   "DB_Integer_S1AHour" : USInt = PLC Data_Integer.S1AHour, 1 s
   "DB_Integer_S1AMinute" : USInt = PLC Data_Integer.S1AMinute, 1 s
   "DB_Integer_S1ASecond" : USInt = PLC Data_Integer.S1ASecond, 1 s
   "DB_Integer_S1BHour" : USInt = PLC Data_Integer.S1BHour, 1 s
   "DB_Integer_S1BMinute" : USInt = PLC Data_Integer.S1BMinute, 1 s
   "DB_Integer_S1BSecond" : USInt = PLC Data_Integer.S1BSecond, 1 s
   "DB_Integer_S2AHour" : USInt = PLC Data_Integer.S2AHour, 1 s
   "DB_Integer_S2AMinute" : USInt = PLC Data_Integer.S2AMinute, 1 s
   "DB_Integer_S2ASecond" : USInt = PLC Data_Integer.S2ASecond, 1 s
   "DB_Integer_S2BHour" : USInt = PLC Data_Integer.S2BHour, 1 s
   "DB_Integer_S2BMinute" : USInt = PLC Data_Integer.S2BMinute, 1 s
   "DB_Integer_S2BSecond" : USInt = PLC Data_Integer.S2BSecond, 1 s
   "DB_Integer_S3AHour" : USInt = PLC Data_Integer.S3AHour, 1 s
   "DB_Integer_S3AMinute" : USInt = PLC Data_Integer.S3AMinute, 1 s
   "DB_Integer_S3ASecond" : USInt = PLC Data_Integer.S3ASecond, 1 s
   "DB_Integer_S3BHour" : USInt = PLC Data_Integer.S3BHour, 1 s
   "DB_Integer_S3BMinute" : USInt = PLC Data_Integer.S3BMinute, 1 s
   "DB_Integer_S3BSecond" : USInt = PLC Data_Integer.S3BSecond, 1 s
   "Data_Bool1_F_Set Time Day" : Bool = PLC Data_Bool1."F_Set Time Day", 1 s
   "Data_integer2_Flag Input Always Bad Read" : USInt = PLC Data_integer2."Flag Input Always Bad Read", 1 s
   "Data_DTLData_DTL_Mesin Run[0].HOUR" : USInt = PLC Data_DTLData."DTL_Mesin Run"[0].HOUR, 1 s
   "Data_DTLData_DTL_Mesin Run[0].MINUTE" : USInt = PLC Data_DTLData."DTL_Mesin Run"[0].MINUTE, 1 s
   "Data_DTLData_DTL_Mesin Run[0].SECOND" : USInt = PLC Data_DTLData."DTL_Mesin Run"[0].SECOND, 1 s
   "Data_Real_%Mesin Run[0]" : Real = PLC Data_Real."%Mesin Run"[0], 1 s
   "Data_DTLData_DTL_Mesin Run Baypass[0].HOUR" : USInt = PLC Data_DTLData."DTL_Mesin Run Baypass"[0].HOUR, 1 s
   "Data_DTLData_DTL_Mesin Run Baypass[0].MINUTE" : USInt = PLC Data_DTLData."DTL_Mesin Run Baypass"[0].MINUTE, 1 s
   "Data_DTLData_DTL_Mesin Run Baypass[0].SECOND" : USInt = PLC Data_DTLData."DTL_Mesin Run Baypass"[0].SECOND, 1 s
   "Data_Real_%Mesin Run Baypass[0]" : Real = PLC Data_Real."%Mesin Run Baypass"[0], 1 s
   "Data_DTLData_DTL_Mesin Stop[0].HOUR" : USInt = PLC Data_DTLData."DTL_Mesin Stop"[0].HOUR, 1 s
   "Data_DTLData_DTL_Mesin Stop[0].MINUTE" : USInt = PLC Data_DTLData."DTL_Mesin Stop"[0].MINUTE, 1 s
   "Data_DTLData_DTL_Mesin Stop[0].SECOND" : USInt = PLC Data_DTLData."DTL_Mesin Stop"[0].SECOND, 1 s
   "Data_Real_%Mesin Stop[0]" : Real = PLC Data_Real."%Mesin Stop"[0], 1 s
   "Data_DTLData_DTL_Mesin Error[0].HOUR" : USInt = PLC Data_DTLData."DTL_Mesin Error"[0].HOUR, 1 s
   "Data_DTLData_DTL_Mesin Error[0].MINUTE" : USInt = PLC Data_DTLData."DTL_Mesin Error"[0].MINUTE, 1 s
   "Data_DTLData_DTL_Mesin Error[0].SECOND" : USInt = PLC Data_DTLData."DTL_Mesin Error"[0].SECOND, 1 s
   "Data_Real_%Mesin Error[0]" : Real = PLC Data_Real."%Mesin Error"[0], 1 s
   "Data_DTLData_DTL_Mesin Run[1].HOUR" : USInt = PLC Data_DTLData."DTL_Mesin Run"[1].HOUR, 1 s
   "Data_DTLData_DTL_Mesin Run[1].MINUTE" : USInt = PLC Data_DTLData."DTL_Mesin Run"[1].MINUTE, 1 s
   "Data_DTLData_DTL_Mesin Run[1].SECOND" : USInt = PLC Data_DTLData."DTL_Mesin Run"[1].SECOND, 1 s
   "Data_Real_%Mesin Run[1]" : Real = PLC Data_Real."%Mesin Run"[1], 1 s
   "Data_DTLData_DTL_Mesin Run Baypass[1].HOUR" : USInt = PLC Data_DTLData."DTL_Mesin Run Baypass"[1].HOUR, 1 s
   "Data_DTLData_DTL_Mesin Run Baypass[1].MINUTE" : USInt = PLC Data_DTLData."DTL_Mesin Run Baypass"[1].MINUTE, 1 s
   "Data_DTLData_DTL_Mesin Run Baypass[1].SECOND" : USInt = PLC Data_DTLData."DTL_Mesin Run Baypass"[1].SECOND, 1 s
   "Data_Real_%Mesin Run Baypass[1]" : Real = PLC Data_Real."%Mesin Run Baypass"[1], 1 s
   "Data_DTLData_DTL_Mesin Stop[1].HOUR" : USInt = PLC Data_DTLData."DTL_Mesin Stop"[1].HOUR, 1 s
   "Data_DTLData_DTL_Mesin Stop[1].MINUTE" : USInt = PLC Data_DTLData."DTL_Mesin Stop"[1].MINUTE, 1 s
   "Data_DTLData_DTL_Mesin Stop[1].SECOND" : USInt = PLC Data_DTLData."DTL_Mesin Stop"[1].SECOND, 1 s
   "Data_Real_%Mesin Stop[1]" : Real = PLC Data_Real."%Mesin Stop"[1], 1 s
   "Data_DTLData_DTL_Mesin Error[1].HOUR" : USInt = PLC Data_DTLData."DTL_Mesin Error"[1].HOUR, 1 s
   "Data_DTLData_DTL_Mesin Error[1].MINUTE" : USInt = PLC Data_DTLData."DTL_Mesin Error"[1].MINUTE, 1 s
   "Data_DTLData_DTL_Mesin Error[1].SECOND" : USInt = PLC Data_DTLData."DTL_Mesin Error"[1].SECOND, 1 s
   "Data_Real_%Mesin Error[1]" : Real = PLC Data_Real."%Mesin Error"[1], 1 s
   "Data_DTLData_DTL_Mesin Run[2].HOUR" : USInt = PLC Data_DTLData."DTL_Mesin Run"[2].HOUR, 1 s
   "Data_DTLData_DTL_Mesin Run[2].MINUTE" : USInt = PLC Data_DTLData."DTL_Mesin Run"[2].MINUTE, 1 s
   "Data_DTLData_DTL_Mesin Run[2].SECOND" : USInt = PLC Data_DTLData."DTL_Mesin Run"[2].SECOND, 1 s
   "Data_Real_%Mesin Run[2]" : Real = PLC Data_Real."%Mesin Run"[2], 1 s
   "Data_DTLData_DTL_Mesin Run Baypass[2].HOUR" : USInt = PLC Data_DTLData."DTL_Mesin Run Baypass"[2].HOUR, 1 s
   "Data_DTLData_DTL_Mesin Run Baypass[2].MINUTE" : USInt = PLC Data_DTLData."DTL_Mesin Run Baypass"[2].MINUTE, 1 s
   "Data_DTLData_DTL_Mesin Run Baypass[2].SECOND" : USInt = PLC Data_DTLData."DTL_Mesin Run Baypass"[2].SECOND, 1 s
   "Data_Real_%Mesin Run Baypass[2]" : Real = PLC Data_Real."%Mesin Run Baypass"[2], 1 s
   "Data_DTLData_DTL_Mesin Stop[2].HOUR" : USInt = PLC Data_DTLData."DTL_Mesin Stop"[2].HOUR, 1 s
   "Data_DTLData_DTL_Mesin Stop[2].MINUTE" : USInt = PLC Data_DTLData."DTL_Mesin Stop"[2].MINUTE, 1 s
   "Data_DTLData_DTL_Mesin Stop[2].SECOND" : USInt = PLC Data_DTLData."DTL_Mesin Stop"[2].SECOND, 1 s
   "Data_Real_%Mesin Stop[2]" : Real = PLC Data_Real."%Mesin Stop"[2], 1 s
   "Data_DTLData_DTL_Mesin Error[2].HOUR" : USInt = PLC Data_DTLData."DTL_Mesin Error"[2].HOUR, 1 s
   "Data_DTLData_DTL_Mesin Error[2].MINUTE" : USInt = PLC Data_DTLData."DTL_Mesin Error"[2].MINUTE, 1 s
   "Data_DTLData_DTL_Mesin Error[2].SECOND" : USInt = PLC Data_DTLData."DTL_Mesin Error"[2].SECOND, 1 s
   "Data_Real_%Mesin Error[2]" : Real = PLC Data_Real."%Mesin Error"[2], 1 s
   "Data_DTLData_DTL_Mesin Run[3].HOUR" : USInt = PLC Data_DTLData."DTL_Mesin Run"[3].HOUR, 1 s
   "Data_DTLData_DTL_Mesin Run[3].MINUTE" : USInt = PLC Data_DTLData."DTL_Mesin Run"[3].MINUTE, 1 s
   "Data_DTLData_DTL_Mesin Run[3].SECOND" : USInt = PLC Data_DTLData."DTL_Mesin Run"[3].SECOND, 1 s
   "Data_Real_%Mesin Run[3]" : Real = PLC Data_Real."%Mesin Run"[3], 1 s
   "Data_DTLData_DTL_Mesin Run Baypass[3].HOUR" : USInt = PLC Data_DTLData."DTL_Mesin Run Baypass"[3].HOUR, 1 s
   "Data_DTLData_DTL_Mesin Run Baypass[3].MINUTE" : USInt = PLC Data_DTLData."DTL_Mesin Run Baypass"[3].MINUTE, 1 s
   "Data_DTLData_DTL_Mesin Run Baypass[3].SECOND" : USInt = PLC Data_DTLData."DTL_Mesin Run Baypass"[3].SECOND, 1 s
   "Data_Real_%Mesin Run Baypass[3]" : Real = PLC Data_Real."%Mesin Run Baypass"[3], 1 s
   "Data_Real_%Mesin Stop[3]" : Real = PLC Data_Real."%Mesin Stop"[3], 1 s
   "Data_Real_%Mesin Error[3]" : Real = PLC Data_Real."%Mesin Error"[3], 1 s
   "Data_DTLData_DTL_Mesin Stop[3].HOUR" : USInt = PLC Data_DTLData."DTL_Mesin Stop"[3].HOUR, 1 s
   "Data_DTLData_DTL_Mesin Stop[3].MINUTE" : USInt = PLC Data_DTLData."DTL_Mesin Stop"[3].MINUTE, 1 s
   "Data_DTLData_DTL_Mesin Stop[3].SECOND" : USInt = PLC Data_DTLData."DTL_Mesin Stop"[3].SECOND, 1 s
   "Data_DTLData_DTL_Mesin Error[3].HOUR" : USInt = PLC Data_DTLData."DTL_Mesin Error"[3].HOUR, 1 s
   "Data_DTLData_DTL_Mesin Error[3].MINUTE" : USInt = PLC Data_DTLData."DTL_Mesin Error"[3].MINUTE, 1 s
   "Data_DTLData_DTL_Mesin Error[3].SECOND" : USInt = PLC Data_DTLData."DTL_Mesin Error"[3].SECOND, 1 s
   "Data_DTLData_DTL_Mesin Run[4].HOUR" : USInt = PLC Data_DTLData."DTL_Mesin Run"[4].HOUR, 1 s
   "Data_DTLData_DTL_Mesin Run[4].MINUTE" : USInt = PLC Data_DTLData."DTL_Mesin Run"[4].MINUTE, 1 s
   "Data_DTLData_DTL_Mesin Run[4].SECOND" : USInt = PLC Data_DTLData."DTL_Mesin Run"[4].SECOND, 1 s
   "Data_Real_%Mesin Run[4]" : Real = PLC Data_Real."%Mesin Run"[4], 1 s
   "Data_Real_%Mesin Run Baypass[4]" : Real = PLC Data_Real."%Mesin Run Baypass"[4], 1 s
   "Data_Real_%Mesin Stop[4]" : Real = PLC Data_Real."%Mesin Stop"[4], 1 s
   "Data_Real_%Mesin Error[4]" : Real = PLC Data_Real."%Mesin Error"[4], 1 s
   "Data_DTLData_DTL_Mesin Run Baypass[4].HOUR" : USInt = PLC Data_DTLData."DTL_Mesin Run Baypass"[4].HOUR, 1 s
   "Data_DTLData_DTL_Mesin Run Baypass[4].MINUTE" : USInt = PLC Data_DTLData."DTL_Mesin Run Baypass"[4].MINUTE, 1 s
   "Data_DTLData_DTL_Mesin Run Baypass[4].SECOND" : USInt = PLC Data_DTLData."DTL_Mesin Run Baypass"[4].SECOND, 1 s
   "Data_DTLData_DTL_Mesin Stop[4].HOUR" : USInt = PLC Data_DTLData."DTL_Mesin Stop"[4].HOUR, 1 s
   "Data_DTLData_DTL_Mesin Stop[4].MINUTE" : USInt = PLC Data_DTLData."DTL_Mesin Stop"[4].MINUTE, 1 s
   "Data_DTLData_DTL_Mesin Stop[4].SECOND" : USInt = PLC Data_DTLData."DTL_Mesin Stop"[4].SECOND, 1 s
   "Data_DTLData_DTL_Mesin Error[4].HOUR" : USInt = PLC Data_DTLData."DTL_Mesin Error"[4].HOUR, 1 s
   "Data_DTLData_DTL_Mesin Error[4].MINUTE" : USInt = PLC Data_DTLData."DTL_Mesin Error"[4].MINUTE, 1 s
   "Data_DTLData_DTL_Mesin Error[4].SECOND" : USInt = PLC Data_DTLData."DTL_Mesin Error"[4].SECOND, 1 s
   "Data_DTLData_DTL_Mesin Run[5].HOUR" : USInt = PLC Data_DTLData."DTL_Mesin Run"[5].HOUR, 1 s
   "Data_DTLData_DTL_Mesin Run[5].MINUTE" : USInt = PLC Data_DTLData."DTL_Mesin Run"[5].MINUTE, 1 s
   "Data_DTLData_DTL_Mesin Run[5].SECOND" : USInt = PLC Data_DTLData."DTL_Mesin Run"[5].SECOND, 1 s
   "Data_Real_%Mesin Run[5]" : Real = PLC Data_Real."%Mesin Run"[5], 1 s
   "Data_Real_%Mesin Run Baypass[5]" : Real = PLC Data_Real."%Mesin Run Baypass"[5], 1 s
   "Data_Real_%Mesin Stop[5]" : Real = PLC Data_Real."%Mesin Stop"[5], 1 s
   "Data_Real_%Mesin Error[5]" : Real = PLC Data_Real."%Mesin Error"[5], 1 s
   "Data_DTLData_DTL_Mesin Run Baypass[5].HOUR" : USInt = PLC Data_DTLData."DTL_Mesin Run Baypass"[5].HOUR, 1 s
   "Data_DTLData_DTL_Mesin Run Baypass[5].MINUTE" : USInt = PLC Data_DTLData."DTL_Mesin Run Baypass"[5].MINUTE, 1 s
   "Data_DTLData_DTL_Mesin Run Baypass[5].SECOND" : USInt = PLC Data_DTLData."DTL_Mesin Run Baypass"[5].SECOND, 1 s
   "Data_DTLData_DTL_Mesin Stop[5].HOUR" : USInt = PLC Data_DTLData."DTL_Mesin Stop"[5].HOUR, 1 s
   "Data_DTLData_DTL_Mesin Stop[5].MINUTE" : USInt = PLC Data_DTLData."DTL_Mesin Stop"[5].MINUTE, 1 s
   "Data_DTLData_DTL_Mesin Stop[5].SECOND" : USInt = PLC Data_DTLData."DTL_Mesin Stop"[5].SECOND, 1 s
   "Data_DTLData_DTL_Mesin Error[5].HOUR" : USInt = PLC Data_DTLData."DTL_Mesin Error"[5].HOUR, 1 s
   "Data_DTLData_DTL_Mesin Error[5].MINUTE" : USInt = PLC Data_DTLData."DTL_Mesin Error"[5].MINUTE, 1 s
   "Data_DTLData_DTL_Mesin Error[5].SECOND" : USInt = PLC Data_DTLData."DTL_Mesin Error"[5].SECOND, 1 s
   "Data_Time_Timer Delay Stamp" : Time = PLC Data_Time."Timer Delay Stamp", 1 s
   "Data_Time_Timer Trigger Barcode" : Time = PLC Data_Time."Timer Trigger Barcode", 1 s
   "Data_Time_Timer Rejector Slof" : Time = PLC Data_Time."Timer Rejector Slof", 1 s
   "Data_Time_Timer AutoReject" : Time = PLC Data_Time."Timer AutoReject", 1 s
   "Data_DTLData_DTL_Always bad Read[0].HOUR" : USInt = PLC Data_DTLData."DTL_Always bad Read"[0].HOUR, 1 s
   "Data_DTLData_DTL_Always bad Read[0].MINUTE" : USInt = PLC Data_DTLData."DTL_Always bad Read"[0].MINUTE, 1 s
   "Data_DTLData_DTL_Always bad Read[0].SECOND" : USInt = PLC Data_DTLData."DTL_Always bad Read"[0].SECOND, 1 s
   "Data_DTLData_DTL_Press Low[0].HOUR" : USInt = PLC Data_DTLData."DTL_Press Low"[0].HOUR, 1 s
   "Data_DTLData_DTL_Press Low[0].MINUTE" : USInt = PLC Data_DTLData."DTL_Press Low"[0].MINUTE, 1 s
   "Data_DTLData_DTL_Press Low[0].SECOND" : USInt = PLC Data_DTLData."DTL_Press Low"[0].SECOND, 1 s
   "Data_DTLData_DTL_Door Open[0].HOUR" : USInt = PLC Data_DTLData."DTL_Door Open"[0].HOUR, 1 s
   "Data_DTLData_DTL_Door Open[0].MINUTE" : USInt = PLC Data_DTLData."DTL_Door Open"[0].MINUTE, 1 s
   "Data_DTLData_DTL_Door Open[0].SECOND" : USInt = PLC Data_DTLData."DTL_Door Open"[0].SECOND, 1 s
   "Data_DTLData_DTL_Total Detail Error[0].HOUR" : USInt = PLC Data_DTLData."DTL_Total Detail Error"[0].HOUR, 1 s
   "Data_DTLData_DTL_Total Detail Error[0].MINUTE" : USInt = PLC Data_DTLData."DTL_Total Detail Error"[0].MINUTE, 1 s
   "Data_DTLData_DTL_Total Detail Error[0].SECOND" : USInt = PLC Data_DTLData."DTL_Total Detail Error"[0].SECOND, 1 s
   "Data_DTLData_DTL_Always bad Read[1].HOUR" : USInt = PLC Data_DTLData."DTL_Always bad Read"[1].HOUR, 1 s
   "Data_DTLData_DTL_Always bad Read[1].MINUTE" : USInt = PLC Data_DTLData."DTL_Always bad Read"[1].MINUTE, 1 s
   "Data_DTLData_DTL_Always bad Read[1].SECOND" : USInt = PLC Data_DTLData."DTL_Always bad Read"[1].SECOND, 1 s
   "Data_DTLData_DTL_Press Low[1].HOUR" : USInt = PLC Data_DTLData."DTL_Press Low"[1].HOUR, 1 s
   "Data_DTLData_DTL_Press Low[1].MINUTE" : USInt = PLC Data_DTLData."DTL_Press Low"[1].MINUTE, 1 s
   "Data_DTLData_DTL_Press Low[1].SECOND" : USInt = PLC Data_DTLData."DTL_Press Low"[1].SECOND, 1 s
   "Data_DTLData_DTL_Door Open[1].HOUR" : USInt = PLC Data_DTLData."DTL_Door Open"[1].HOUR, 1 s
   "Data_DTLData_DTL_Door Open[1].MINUTE" : USInt = PLC Data_DTLData."DTL_Door Open"[1].MINUTE, 1 s
   "Data_DTLData_DTL_Door Open[1].SECOND" : USInt = PLC Data_DTLData."DTL_Door Open"[1].SECOND, 1 s
   "Data_DTLData_DTL_Always bad Read[2].HOUR" : USInt = PLC Data_DTLData."DTL_Always bad Read"[2].HOUR, 1 s
   "Data_DTLData_DTL_Always bad Read[2].MINUTE" : USInt = PLC Data_DTLData."DTL_Always bad Read"[2].MINUTE, 1 s
   "Data_DTLData_DTL_Always bad Read[2].SECOND" : USInt = PLC Data_DTLData."DTL_Always bad Read"[2].SECOND, 1 s
   "Data_DTLData_DTL_Press Low[2].HOUR" : USInt = PLC Data_DTLData."DTL_Press Low"[2].HOUR, 1 s
   "Data_DTLData_DTL_Press Low[2].MINUTE" : USInt = PLC Data_DTLData."DTL_Press Low"[2].MINUTE, 1 s
   "Data_DTLData_DTL_Press Low[2].SECOND" : USInt = PLC Data_DTLData."DTL_Press Low"[2].SECOND, 1 s
   "Data_DTLData_DTL_Door Open[2].HOUR" : USInt = PLC Data_DTLData."DTL_Door Open"[2].HOUR, 1 s
   "Data_DTLData_DTL_Door Open[2].MINUTE" : USInt = PLC Data_DTLData."DTL_Door Open"[2].MINUTE, 1 s
   "Data_DTLData_DTL_Door Open[2].SECOND" : USInt = PLC Data_DTLData."DTL_Door Open"[2].SECOND, 1 s
   "Data_DTLData_DTL_Always bad Read[3].HOUR" : USInt = PLC Data_DTLData."DTL_Always bad Read"[3].HOUR, 1 s
   "Data_DTLData_DTL_Always bad Read[3].MINUTE" : USInt = PLC Data_DTLData."DTL_Always bad Read"[3].MINUTE, 1 s
   "Data_DTLData_DTL_Always bad Read[3].SECOND" : USInt = PLC Data_DTLData."DTL_Always bad Read"[3].SECOND, 1 s
   "Data_DTLData_DTL_Press Low[3].HOUR" : USInt = PLC Data_DTLData."DTL_Press Low"[3].HOUR, 1 s
   "Data_DTLData_DTL_Press Low[3].MINUTE" : USInt = PLC Data_DTLData."DTL_Press Low"[3].MINUTE, 1 s
   "Data_DTLData_DTL_Press Low[3].SECOND" : USInt = PLC Data_DTLData."DTL_Press Low"[3].SECOND, 1 s
   "Data_DTLData_DTL_Door Open[3].HOUR" : USInt = PLC Data_DTLData."DTL_Door Open"[3].HOUR, 1 s
   "Data_DTLData_DTL_Door Open[3].MINUTE" : USInt = PLC Data_DTLData."DTL_Door Open"[3].MINUTE, 1 s
   "Data_DTLData_DTL_Door Open[3].SECOND" : USInt = PLC Data_DTLData."DTL_Door Open"[3].SECOND, 1 s
   "Data_DTLData_DTL_Always bad Read[4].HOUR" : USInt = PLC Data_DTLData."DTL_Always bad Read"[4].HOUR, 1 s
   "Data_DTLData_DTL_Always bad Read[4].MINUTE" : USInt = PLC Data_DTLData."DTL_Always bad Read"[4].MINUTE, 1 s
   "Data_DTLData_DTL_Always bad Read[4].SECOND" : USInt = PLC Data_DTLData."DTL_Always bad Read"[4].SECOND, 1 s
   "Data_DTLData_DTL_Press Low[4].HOUR" : USInt = PLC Data_DTLData."DTL_Press Low"[4].HOUR, 1 s
   "Data_DTLData_DTL_Press Low[4].MINUTE" : USInt = PLC Data_DTLData."DTL_Press Low"[4].MINUTE, 1 s
   "Data_DTLData_DTL_Press Low[4].SECOND" : USInt = PLC Data_DTLData."DTL_Press Low"[4].SECOND, 1 s
   "Data_DTLData_DTL_Door Open[4].HOUR" : USInt = PLC Data_DTLData."DTL_Door Open"[4].HOUR, 1 s
   "Data_DTLData_DTL_Door Open[4].MINUTE" : USInt = PLC Data_DTLData."DTL_Door Open"[4].MINUTE, 1 s
   "Data_DTLData_DTL_Door Open[4].SECOND" : USInt = PLC Data_DTLData."DTL_Door Open"[4].SECOND, 1 s
   "Data_DTLData_DTL_Always bad Read[5].HOUR" : USInt = PLC Data_DTLData."DTL_Always bad Read"[5].HOUR, 1 s
   "Data_DTLData_DTL_Always bad Read[5].MINUTE" : USInt = PLC Data_DTLData."DTL_Always bad Read"[5].MINUTE, 1 s
   "Data_DTLData_DTL_Always bad Read[5].SECOND" : USInt = PLC Data_DTLData."DTL_Always bad Read"[5].SECOND, 1 s
   "Data_DTLData_DTL_Press Low[5].HOUR" : USInt = PLC Data_DTLData."DTL_Press Low"[5].HOUR, 1 s
   "Data_DTLData_DTL_Press Low[5].MINUTE" : USInt = PLC Data_DTLData."DTL_Press Low"[5].MINUTE, 1 s
   "Data_DTLData_DTL_Press Low[5].SECOND" : USInt = PLC Data_DTLData."DTL_Press Low"[5].SECOND, 1 s
   "Data_DTLData_DTL_Door Open[5].HOUR" : USInt = PLC Data_DTLData."DTL_Door Open"[5].HOUR, 1 s
   "Data_DTLData_DTL_Door Open[5].MINUTE" : USInt = PLC Data_DTLData."DTL_Door Open"[5].MINUTE, 1 s
   "Data_DTLData_DTL_Door Open[5].SECOND" : USInt = PLC Data_DTLData."DTL_Door Open"[5].SECOND, 1 s
   "Data_IntData_Label Sloft[0]" : UDInt = PLC Data_IntData."Label Sloft"[0], 1 s
   "Data_IntData_Un label Sloft[0]" : UDInt = PLC Data_IntData."Un label Sloft"[0], 1 s
   "Data_IntData_Label Sloft[1]" : UDInt = PLC Data_IntData."Label Sloft"[1], 1 s
   "Data_IntData_Un label Sloft[1]" : UDInt = PLC Data_IntData."Un label Sloft"[1], 1 s
   "Data_IntData_Label Sloft[2]" : UDInt = PLC Data_IntData."Label Sloft"[2], 1 s
   "Data_IntData_Un label Sloft[2]" : UDInt = PLC Data_IntData."Un label Sloft"[2], 1 s
   "Data_IntData_Label Sloft[3]" : UDInt = PLC Data_IntData."Label Sloft"[3], 1 s
   "Data_IntData_Un label Sloft[3]" : UDInt = PLC Data_IntData."Un label Sloft"[3], 1 s
   "Data_IntData_Label Sloft[4]" : UDInt = PLC Data_IntData."Label Sloft"[4], 1 s
   "Data_IntData_Un label Sloft[4]" : UDInt = PLC Data_IntData."Un label Sloft"[4], 1 s
   "Data_IntData_Label Sloft[5]" : UDInt = PLC Data_IntData."Label Sloft"[5], 1 s
   "Data_IntData_Un label Sloft[5]" : UDInt = PLC Data_IntData."Un label Sloft"[5], 1 s
   "Data_Real_% label Sloft[0]" : Real = PLC Data_Real."% label Sloft"[0], 1 s
   "Data_Real_% Unlabel Sloft[0]" : Real = PLC Data_Real."% Unlabel Sloft"[0], 1 s
   "Data_Real_% label Sloft[1]" : Real = PLC Data_Real."% label Sloft"[1], 1 s
   "Data_Real_% Unlabel Sloft[1]" : Real = PLC Data_Real."% Unlabel Sloft"[1], 1 s
   "Data_Real_% label Sloft[2]" : Real = PLC Data_Real."% label Sloft"[2], 1 s
   "Data_Real_% Unlabel Sloft[2]" : Real = PLC Data_Real."% Unlabel Sloft"[2], 1 s
   "Data_Real_% label Sloft[3]" : Real = PLC Data_Real."% label Sloft"[3], 1 s
   "Data_Real_% Unlabel Sloft[3]" : Real = PLC Data_Real."% Unlabel Sloft"[3], 1 s
   "Data_Real_% label Sloft[4]" : Real = PLC Data_Real."% label Sloft"[4], 1 s
   "Data_Real_% Unlabel Sloft[4]" : Real = PLC Data_Real."% Unlabel Sloft"[4], 1 s
   "Data_Real_% label Sloft[5]" : Real = PLC Data_Real."% label Sloft"[5], 1 s
   "Data_Real_% Unlabel Sloft[5]" : Real = PLC Data_Real."% Unlabel Sloft"[5], 1 s
   "Data_IntData_Sloft Bypass[0]" : UDInt = PLC Data_IntData."Sloft Bypass"[0], 1 s
   "Data_IntData_Sloft Bypass[1]" : UDInt = PLC Data_IntData."Sloft Bypass"[1], 1 s
   "Data_IntData_Sloft Bypass[2]" : UDInt = PLC Data_IntData."Sloft Bypass"[2], 1 s
   "Data_IntData_Sloft Bypass[3]" : UDInt = PLC Data_IntData."Sloft Bypass"[3], 1 s
   "Data_IntData_Sloft Bypass[4]" : UDInt = PLC Data_IntData."Sloft Bypass"[4], 1 s
   "Data_IntData_Sloft Bypass[5]" : UDInt = PLC Data_IntData."Sloft Bypass"[5], 1 s
   "Data_Real_% Sloft bypass[0]" : Real = PLC Data_Real."% Sloft bypass"[0], 1 s
   "Data_Real_% Sloft bypass[1]" : Real = PLC Data_Real."% Sloft bypass"[1], 1 s
   "Data_Real_% Sloft bypass[2]" : Real = PLC Data_Real."% Sloft bypass"[2], 1 s
   "Data_Real_% Sloft bypass[3]" : Real = PLC Data_Real."% Sloft bypass"[3], 1 s
   "Data_Real_% Sloft bypass[4]" : Real = PLC Data_Real."% Sloft bypass"[4], 1 s
   "Data_Real_% Sloft bypass[5]" : Real = PLC Data_Real."% Sloft bypass"[5], 1 s
   "Data_IntData_uintDT_AplicatorFreeze[0]" : UInt = PLC Data_IntData.uintDT_AplicatorFreeze[0], 1 s
   "Data_IntData_uintDT_AplicatorFreeze[1]" : UInt = PLC Data_IntData.uintDT_AplicatorFreeze[1], 1 s
   "Data_IntData_uintDT_AplicatorFreeze[2]" : UInt = PLC Data_IntData.uintDT_AplicatorFreeze[2], 1 s
   "Data_IntData_uintDT_AplicatorFreeze[3]" : UInt = PLC Data_IntData.uintDT_AplicatorFreeze[3], 1 s
   "Data_IntData_uintDT_AplicatorFreeze[4]" : UInt = PLC Data_IntData.uintDT_AplicatorFreeze[4], 1 s
   "Data_IntData_uintDT_AplicatorFreeze[5]" : UInt = PLC Data_IntData.uintDT_AplicatorFreeze[5], 1 s
   "Data_DTLData_Total Time Machine[0].HOUR" : USInt = PLC Data_DTLData."Total Time Machine"[0].HOUR, 1 s
   "Data_DTLData_Total Time Machine[0].MINUTE" : USInt = PLC Data_DTLData."Total Time Machine"[0].MINUTE, 1 s
   "Data_DTLData_Total Time Machine[0].SECOND" : USInt = PLC Data_DTLData."Total Time Machine"[0].SECOND, 1 s
   "Data_DTLData_Total Time Machine[1].HOUR" : USInt = PLC Data_DTLData."Total Time Machine"[1].HOUR, 1 s
   "Data_DTLData_Total Time Machine[1].MINUTE" : USInt = PLC Data_DTLData."Total Time Machine"[1].MINUTE, 1 s
   "Data_DTLData_Total Time Machine[1].SECOND" : USInt = PLC Data_DTLData."Total Time Machine"[1].SECOND, 1 s
   "Data_DTLData_Total Time Machine[2].HOUR" : USInt = PLC Data_DTLData."Total Time Machine"[2].HOUR, 1 s
   "Data_DTLData_Total Time Machine[2].MINUTE" : USInt = PLC Data_DTLData."Total Time Machine"[2].MINUTE, 1 s
   "Data_DTLData_Total Time Machine[2].SECOND" : USInt = PLC Data_DTLData."Total Time Machine"[2].SECOND, 1 s
   "Data_DTLData_Total Time Machine[3].HOUR" : USInt = PLC Data_DTLData."Total Time Machine"[3].HOUR, 1 s
   "Data_DTLData_Total Time Machine[3].MINUTE" : USInt = PLC Data_DTLData."Total Time Machine"[3].MINUTE, 1 s
   "Data_DTLData_Total Time Machine[3].SECOND" : USInt = PLC Data_DTLData."Total Time Machine"[3].SECOND, 1 s
   "Data_DTLData_Total Time Machine[4].HOUR" : USInt = PLC Data_DTLData."Total Time Machine"[4].HOUR, 1 s
   "Data_DTLData_Total Time Machine[4].MINUTE" : USInt = PLC Data_DTLData."Total Time Machine"[4].MINUTE, 1 s
   "Data_DTLData_Total Time Machine[4].SECOND" : USInt = PLC Data_DTLData."Total Time Machine"[4].SECOND, 1 s
   "Data_DTLData_Total Time Machine[5].HOUR" : USInt = PLC Data_DTLData."Total Time Machine"[5].HOUR, 1 s
   "Data_DTLData_Total Time Machine[5].MINUTE" : USInt = PLC Data_DTLData."Total Time Machine"[5].MINUTE, 1 s
   "Data_DTLData_Total Time Machine[5].SECOND" : USInt = PLC Data_DTLData."Total Time Machine"[5].SECOND, 1 s
   "Data_DTLData_DTL_Total Detail Error[5].HOUR" : USInt = PLC Data_DTLData."DTL_Total Detail Error"[5].HOUR, 1 s
   "Data_DTLData_DTL_Total Detail Error[5].MINUTE" : USInt = PLC Data_DTLData."DTL_Total Detail Error"[5].MINUTE, 1 s
   "Data_DTLData_DTL_Total Detail Error[5].SECOND" : USInt = PLC Data_DTLData."DTL_Total Detail Error"[5].SECOND, 1 s
   "Data_DTLData_DTL_Total Detail Error[4].HOUR" : USInt = PLC Data_DTLData."DTL_Total Detail Error"[4].HOUR, 1 s
   "Data_DTLData_DTL_Total Detail Error[4].MINUTE" : USInt = PLC Data_DTLData."DTL_Total Detail Error"[4].MINUTE, 1 s
   "Data_DTLData_DTL_Total Detail Error[4].SECOND" : USInt = PLC Data_DTLData."DTL_Total Detail Error"[4].SECOND, 1 s
   "Data_DTLData_DTL_Total Detail Error[3].HOUR" : USInt = PLC Data_DTLData."DTL_Total Detail Error"[3].HOUR, 1 s
   "Data_DTLData_DTL_Total Detail Error[3].MINUTE" : USInt = PLC Data_DTLData."DTL_Total Detail Error"[3].MINUTE, 1 s
   "Data_DTLData_DTL_Total Detail Error[3].SECOND" : USInt = PLC Data_DTLData."DTL_Total Detail Error"[3].SECOND, 1 s
   "Data_DTLData_DTL_Total Detail Error[2].HOUR" : USInt = PLC Data_DTLData."DTL_Total Detail Error"[2].HOUR, 1 s
   "Data_DTLData_DTL_Total Detail Error[2].MINUTE" : USInt = PLC Data_DTLData."DTL_Total Detail Error"[2].MINUTE, 1 s
   "Data_DTLData_DTL_Total Detail Error[2].SECOND" : USInt = PLC Data_DTLData."DTL_Total Detail Error"[2].SECOND, 1 s
   "Data_DTLData_DTL_Total Detail Error[1].HOUR" : USInt = PLC Data_DTLData."DTL_Total Detail Error"[1].HOUR, 1 s
   "Data_DTLData_DTL_Total Detail Error[1].MINUTE" : USInt = PLC Data_DTLData."DTL_Total Detail Error"[1].MINUTE, 1 s
   "Data_DTLData_DTL_Total Detail Error[1].SECOND" : USInt = PLC Data_DTLData."DTL_Total Detail Error"[1].SECOND, 1 s
   "Data_String_sDT_Machine id" : String[254] = PLC Data_String."sDT_Machine id", 1 s
   "RS_Bypass_Addrej" : Bool = PLC RS_Bypass_Addrej AT %M31.4, 1 s
   "Data_IntData_InReject" : UDInt = PLC Data_IntData.InReject, 1 s
   "Data_IntData_InReject_1" : UDInt = PLC Data_IntData.InReject_1, 1 s
   "Data_IntData_InReject_2" : UDInt = PLC Data_IntData.InReject_2, 1 s
   "Data_IntData_InReject_3" : UDInt = PLC Data_IntData.InReject_3, 1 s
   "Data_IntData_InReject_4" : UDInt = PLC Data_IntData.InReject_4, 1 s
   "Data_IntData_InReject_5" : UDInt = PLC Data_IntData.InReject_5, 1 s
   "Data_Real_%InputReject[5]" : Real = PLC Data_Real.%InputReject[5], 1 s
   "Data_Real_%InputReject[4]" : Real = PLC Data_Real.%InputReject[4], 1 s
   "Data_Real_%InputReject[3]" : Real = PLC Data_Real.%InputReject[3], 1 s
   "Data_Real_%InputReject[2]" : Real = PLC Data_Real.%InputReject[2], 1 s
   "Data_Real_%InputReject[1]" : Real = PLC Data_Real.%InputReject[1], 1 s
   "Data_Real_%InputReject[0]" : Real = PLC Data_Real.%InputReject[0], 1 s
   "AddReject2_DB_Countaddrej" : Time = PLC AddReject2_DB.Countaddrej, 1 s
   "AddReject2_DB_CountStop" : Bool = PLC AddReject2_DB.CountStop, 1 s

discrete alarms
   1: 'Pressure Low', class Errors, trigger "HMI_Tag_1" bit 8
   2: 'Door Open Labelling', class Errors, trigger "HMI_Tag_1" bit 9
   3: 'Door Open Focke Chute', class Errors, trigger "HMI_Tag_1" bit 10
   4: 'Chute 3 Way Full', class Errors, trigger "HMI_Tag_1" bit 11
   5: 'Door Open FC Proximity', class Errors, trigger "HMI_Tag_1" bit 12
   6: 'Alarm2', class Errors, trigger "HMI_Tag_1" bit 13
   7: 'Imaje Paper/Ribbon Out', class Errors, trigger "HMI_Tag_1" bit 14
   8: 'Imaje System Error', class Errors, trigger "HMI_Tag_1" bit 15
   9: 'Imaje Not In Position', class Errors, trigger "HMI_Tag_1" bit 0
   10: 'Heater Not Ready', class Errors, trigger "HMI_Tag_1" bit 1
   11: 'Reed Switch Pneumatic 1 Pusher', class Errors, trigger "HMI_Tag_1" bit 2
   12: 'Reed Switch Pneumatic 1 Pusher Retract', class Errors, trigger "HMI_Tag_1" bit 3
   13: 'Reed Switch Pneumatic 3 Up', class Errors, trigger "HMI_Tag_1" bit 4
   14: 'Reed Switch Pneumatic 3 Down', class Errors, trigger "HMI_Tag_1" bit 5
   15: 'Reed Switch Pneumatic 4 Down', class Errors, trigger "HMI_Error_Cont" bit 8
   16: 'Reed Switch Pneumatic 4 Up', class Errors, trigger "HMI_Error_Cont" bit 9
   17: 'Reed Switch Pneumatic 5 Advance', class Errors, trigger "HMI_Error_Cont" bit 10
   18: 'Reed Switch Pneumatic 5 Retract', class Errors, trigger "HMI_Error_Cont" bit 11
   19: 'Chute Heating Roll Full', class Errors, trigger "HMI_Tag_1" bit 6
   20: 'Conveyor Outfeed jammed', class Errors, trigger "HMI_Error_Cont" bit 12
   21: 'Sloft Jammed', class Errors, trigger "HMI_Error_Cont" bit 13
   22: 'Sloft Jammed Infeed Chute', class Errors, trigger "HMI_Error_Cont" bit 14
   24: 'Always Bad Read Sloft', class Errors, trigger "HMI_Error_Cont" bit 15
   23: 'Paper Or Ribbon Low', class Errors, trigger "HMI_Error_Cont" bit 0
   25: 'Emergency Stop Push', class Errors, trigger "HMI_Error_Cont" bit 1

text list "Machine Running": 0 'STOP'; 1 'RUNNING'

text list "Status Markem": 0 'PAUSE'; 1 'START'

text list "Mode Machine": 0 'With Focke Chute'; 1 'Without Focke Chute'

text list "Mode Bypass": 0 'OFF'; 1 'ON'

Template "Template_1" 320x240
   Button "Template_" at 267,190 size 51x47; TextOff 'ExitRuntime'; PictureOff "ExitRuntime_HMI_1"; PictureOn "ExitRuntime_HMI_1"
      on Release: StopRuntime(0)
   Button "Template_1" at 214,190 size 51x47; TextOff 'Text'
   Button "Template_2" at 160,190 size 51x47; TextOff 'Text'
   Button "Template_3" at 107,190 size 51x47; TextOff 'Login'; PictureOff "Login_HMI_1"; PictureOn "Login_HMI_1"
      on Release: function_a2a04561()
   Button "Template_4" at 54,190 size 51x47; TextOff 'AlarmDisplay'; PictureOff "AlarmDisplay_HMI_1"; PictureOn "AlarmDisplay_HMI_1"
      on Release: function_ef3f5d25("Alarm window_Unacknowledged", -1)
   Button "Template_5" at 1,190 size 51x47; TextOff 'NavigateHome'; PictureOff "NavigateHome_HMI_1"; PictureOn "NavigateHome_HMI_1"
   SymbolicIOField "Symbolic_IO_Field_Screen" at 73,7 size 160x25; TextOff '0'; TextOn '1'; TextList "TextList_ScreenNames"
      ProcessValue <- "Tag_ScreenNumber"
   DateTimeField "Template_6" at 235,20 size 85x20
   DateTimeField "Template_7" at 235,0 size 85x20
   GraphicView "Logo" at 0,0 size 71x40; Picture "Logo of HMI_1"

screen "Introduction" 320x240
   Button "Button_1" at 100,200 size 120x30; TextOff 'Go to Main Page'
      on Click: ActivateScreen("Main Page", 0)
   GraphicView "Graphic view_1" at 0,0 size 319x37; Picture "Logo SMS"
   TextField "Text field_1" at 6,54 size 278x31; Text 'END LABELLER MACHINE'
   Button "Button_2" at 7,37 size 29x24; TextOff 'Door Open Secret'
      on Click: ActivateScreen("Door Open Secret", 0)
   TextField "Text field_3" at 20,73 size 278x88; Text 'Compressed Air : 6 Bar Year : 2014 Program Version : 14.06.02'

screen "Main Page" 320x240
   on GenerateScreen: SetBit("Flag Main Page")
   TextField "Text field_1" at 106,1 size 113x25; Text 'MAIN PAGE'
   TextField "Text field_3" at 5,64 size 91x15; Text 'Machine Status'
   TextField "Text field_4" at 5,87 size 91x15; Text 'Markem Status'
   SymbolicIOField "Symbolic I/O field_2" at 100,62 size 122x19; TextOff '0'; TextOn '1'; TextList "Machine Running"
      ProcessValue <- "Machine Running"
   SymbolicIOField "Symbolic I/O field_1" at 100,85 size 122x19; TextOff '0'; TextOn '1'; TextList "Status Markem"
      ProcessValue <- "Flag Imaje Start"
   Button "Button_4" at 0,209 size 90x30; TextOff 'Test Mode'
      on Click: ActivateScreen("Test Mode", 0)
   Button "Button_5" at 95,209 size 90x30; TextOff 'Parameter'
      on Click: ActivateScreen("Parameter", 0)
   TextField "Text field_5" at 5,109 size 91x15; Text 'Mode Machine'
   SymbolicIOField "Symbolic I/O field_3" at 100,108 size 122x19; TextOff '0'; TextOn '1'; TextList "Mode Machine"
      ProcessValue <- "Flag Enable/Disable Block Focke"
   TextField "Text field_7" at 5,131 size 91x15; Text 'Mode Bypass'
   SymbolicIOField "Symbolic I/O field_4" at 100,131 size 122x19; TextOff '0'; TextOn '1'; TextList "Mode Bypass"
      ProcessValue <- "Flag Machine Bypass"
   Button "Button_1" at 289,1 size 29x24; TextOff 'Text'
      on Press: StopRuntime(0)
   IOField "I/O field_3" at 84,26 size 155x23; FormatPattern 9999999999999999999999999999999999999999
      ProcessValue <- "Data_DTL1_Output"
   Button "Button_2" at 191,209 size 103x30; TextOff 'Statistic Data'; TextOn 'Statistika Data'
      on Click: ActivateScreen("St_Data Statistic", 0)
   IOField "I/O field_1" at 124,41 size 76x17; FormatPattern ????????
      ProcessValue <- "Data_String_sDT_Machine id"

screen "Parameter" 320x240
   on GenerateScreen: SetBit("Flag Parameter Page")
   on ClearScreen: ResetBit("Flag Parameter Page")
   TextField "Text field_1" at 1,0 size 319x27; Text 'PARAMETER'
   Button "Button_4" at 91,202 size 132x30; TextOff 'Back to Main Page'
      on Click: ActivateScreen("Main Page", 0)
   Button "Button_3" at 91,48 size 132x30; TextOff 'Setting Timer And Data'; TextOn 'Setting Timer'
      on Click: ActivateScreen("Setting Timer", 0)
   Button "Button_2" at 91,88 size 132x30; TextOff 'Setting Machine'
      on Click: ActivateScreen("Setting Machine", 0)

screen "Setting Timer" 320x240
   on ClearScreen: ResetBit("Flag Parameter Page")
   on GenerateScreen: SetBit("Flag Parameter Page")
   TextField "Text field_1" at 0,0 size 319x27; Text 'SETTING TIMER'
   Button "Button_2" at 92,200 size 120x30; TextOff 'Back to Parameter'
      on Click: ActivateScreen("Parameter", 0)
   TextField "Text field_2" at 1,39 size 150x15; Text 'Timer Delay Stamp'
   IOField "I/O field_1" at 152,40 size 80x16; FormatPattern 9999; Unit  ms
      ProcessValue <- "Data_Time_Timer Delay Stamp"
   TextField "Text field_3" at 2,63 size 150x15; Text 'Timer Trigger Barcode'
   IOField "I/O field_2" at 152,64 size 80x16; FormatPattern 9999; Unit  ms
      ProcessValue <- "Data_Time_Timer Trigger Barcode"
   TextField "Text field_4" at 10,88 size 142x15; Text 'Timer Rejector'
   IOField "I/O field_3" at 152,88 size 80x16; FormatPattern 9999; Unit  ms
      ProcessValue <- "Data_Time_Timer Rejector Slof"
   IOField "I/O field_4" at 152,112 size 80x16; FormatPattern 9999; Unit  ms
      ProcessValue <- "Data_Time_Timer AutoReject"
   TextField "Text field_5" at 8,112 size 142x15; Text 'Timer AutoReject Outfeed'
   TextField "Text field_7" at 5,149 size 143x15; Text 'Total Value Always Bad Read'
   IOField "I/O field_6" at 151,149 size 80x16; FormatPattern 999; Unit  pcs
      ProcessValue <- "Data_integer2_Flag Input Always Bad Read"
   TextField "Text field_8" at 7,172 size 140x15; Text 'Machine Id (Max 8 Char)'
   IOField "I/O field_7" at 152,172 size 81x16; FormatPattern ????????
      ProcessValue <- "Data_String_sDT_Machine id"

screen "Test Mode" 320x240
   on GenerateScreen: SetBit("PB Test Mode")
   on ClearScreen: ResetBit("PB Test Mode")
   TextField "Text field_1" at 1,1 size 319x27; Text 'TEST MODE'
   Switch "Switch_1" at 3,34 size 95x30; TextOff 'Pneumatic 1 Off'; CaptionText 'Switch'; TextOn 'Pneumatic 1 On'
      ProcessValue <- "PB Test Pneumatic 1"
   Switch "Switch_2" at 3,75 size 95x30; CaptionText 'Switch'; TextOff 'Pneumatic 2 Off'; TextOn 'Pneumatic 2 On'
      ProcessValue <- "PB Test Pneumatic 2"
   Switch "Switch_3" at 3,116 size 95x30; CaptionText 'Switch'; TextOff 'Pneumatic 3 Off'; TextOn 'Pneumatic 3 On'
      ProcessValue <- "PB Test Pneumatic 3"
   Switch "Switch_5" at 104,34 size 115x30; CaptionText 'Switch'; TextOff 'Pneumatic 5 Off'; TextOn 'Pneumatic 5 On'
      ProcessValue <- "PB Test Pneumatic 5"
   Switch "Switch_6" at 226,116 size 90x30; CaptionText 'Switch'; TextOff 'Motor Off'; TextOn 'Motor On'
      ProcessValue <- "PB Test Motor"
   Button "Button_1" at 100,204 size 120x30; TextOff 'Back to Main Page'
      on Click: ActivateScreen("Main Page", 0)
   Button "Button_2" at 226,34 size 90x30; TextOff 'Stamp Off'; TextOn 'Stamp On'
      on Press: SetBit("PB Test Imaje")
      on Release: ResetBit("PB Test Imaje")
   Switch "Switch_7" at 104,116 size 115x30; CaptionText 'Switch'; TextOff 'Air Valve On'; TextOn 'Air Valve Off'
      ProcessValue <- "PB Test Air Valve"
   Button "Button_3" at 226,75 size 90x30; TextOff 'Teach In'
      on Press: SetBit("Flag Teach In Barcode")
      on Release: ResetBit("Flag Teach In Barcode")
   Switch "Switch_8" at 3,157 size 95x30; CaptionText 'Switch'; TextOff 'Pneumatic 4 Off'; TextOn 'Pneumatic 4 On'
      ProcessValue <- "PB Test Pneumatic 4"
   Switch "Switch_4" at 104,75 size 115x30; CaptionText 'Switch'; TextOff 'Pneumatic 6 On'; TextOn 'Pneumatic 6 Off'
      ProcessValue <- "PB Test Pneumatic 6"
   Switch "Switch_9" at 104,157 size 115x30; CaptionText 'Switch'; TextOff 'Conveyor Pusher Off'; TextOn 'Conveyor Pusher On'
      ProcessValue <- "PB Test Motor Coveyor Pusher"

screen "Setting Machine" 320x240
   on ClearScreen: ResetBit("Flag Parameter Page")
   on GenerateScreen: SetBit("Flag Parameter Page")
   TextField "Text field_1" at 1,0 size 319x27; Text 'SETTING MACHINE'
   Switch "Switch_1" at 16,38 size 135x30; CaptionText 'Switch'; TextOff 'Barcode ON'; TextOn 'Barcode Off'
      ProcessValue <- "Flag Barcode HMI"
   Switch "Switch_2" at 16,73 size 135x30; CaptionText 'Switch'; TextOff 'Chute 3Way Error ON'; TextOn 'Chute 3Way Error OFF'
      ProcessValue <- "Flag Enable/Disable Error Chute 3 Way"
   Button "Button_2" at 101,205 size 120x30; TextOff 'Back to Parameter'
      on Click: ActivateScreen("Parameter", 0)
   Switch "Switch_4" at 170,38 size 135x30; CaptionText 'Switch'; TextOff 'Reed Switch Bypass Off'; TextOn 'Reed Switch Bypass On'
      ProcessValue <- "Flag Pneumatic Bypass"
   Button "Button_1" at 289,0 size 31x30; TextOff 'Setting Mode'; Authorization "User administration"
      on Click: ActivateScreen("Setting Mode", 0)
   Button "Button_3" at 170,73 size 135x30; TextOff 'Setting Reed Switch'
      on Click: ActivateScreen("Setting Reed Switch", 0)
   Softkey "Softkey_F6" at 266,202 size 53x38
      on KeyDown: ActivateScreen("Setting Mode", 0)
      on KeyUp: ActivateScreen("Setting Mode", 0)
   Softkey "Softkey_F5" at 213,202 size 53x38
      on KeyDown: function_f23ef4c9()
      on KeyUp: function_f23ef4c9()

screen "Setting Mode" 320x240
   TextField "Text field_1" at 1,0 size 319x27; Text 'MODE MACHINE'
   Button "Button_1" at 95,203 size 129x30; TextOff 'Back to Setting Machine'
      on Click: ActivateScreen("Setting Machine", 0)
   Switch "Switch_1" at 69,36 size 177x32; CaptionText 'Switch'; TextOff 'With Focke Chute'; TextOn 'Without Focke Chute'
      ProcessValue <- "Flag Enable/Disable Block Focke"
   Switch "Switch_2" at 69,71 size 177x32; TextOff 'Disable Reject Markem Error'; CaptionText 'Switch'; TextOn 'Enable Reject Markem Error'
      ProcessValue <- "Flag Enable/Disable Flow to Reject"
   Switch "Switch_3" at 69,108 size 177x32; TextOff 'Enable Reject Outfeed Stop'; CaptionText 'Switch'; TextOn 'Disable Reject Outfeed Stop'
      ProcessValue <- "Flag Enable/Disable Reject Outfeed"

screen "Setting Reed Switch" 320x240
   TextField "Text field_1" at 1,3 size 319x27; Text 'SETTING REED SWITCH BYPASS'
   Switch "Switch_4" at 21,103 size 128x30; CaptionText 'Switch'; TextOff 'RS Pneu 3 Bypass Off'; TextOn 'RS Pneu 3 Bypass On'
      ProcessValue <- "RS Bypass Pneumatic 3"
   Switch "Switch_1" at 172,103 size 128x30; CaptionText 'Switch'; TextOff 'RS Pneu 5 Bypass Off'; TextOn 'RS Pneu 5 Bypass On'
      ProcessValue <- "RS Bypass Pneumatic 5"
   Switch "Switch_2" at 172,59 size 128x30; CaptionText 'Switch'; TextOff 'RS Pneu 4 Bypass Off'; TextOn 'RS Pneu 4 Bypass On'
      ProcessValue <- "RS Bypass Pneumatic 4"
   Switch "Switch_3" at 21,59 size 128x30; CaptionText 'Switch'; TextOff 'RS Pneu 1 Bypass Off'; TextOn 'RS Pneu 1 Bypass On'
      ProcessValue <- "RS Bypass Pneumatic 1"
   Button "Button_1" at 95,203 size 129x30; TextOff 'Back to Setting Machine'
      on Click: ActivateScreen("Setting Machine", 0)
   Switch "Switch_5" at 172,143 size 128x30; TextOff 'RS Pneu 7 Bypass Off'; TextOn 'RS Pneu 7 Bypass On'; CaptionText 'Switch'
      ProcessValue <- "RS_Bypass_Addrej"

screen "St_Data Statistic" 320x240
   Button "Button_1" at 9,47 size 146x30; TextOff 'Current Shift Data'
      on Click: ActivateScreen("St_Quantity Data", 0)
   Button "Button_2" at 287,3 size 27x24; TextOff 'Text'; TextOn 'Statistik Parameter'; Authorization "User administration"
      on Click: ActivateScreen("St_Parameter", 0)
   Button "Button_3" at 9,80 size 146x30; TextOff 'Current Shift Data Minus 1'
      on Click: ActivateScreen("St_Quantity Data_1", 0)
   Button "Button_4" at 9,113 size 147x30; TextOff 'Current Shift Data Minus 2'
      on Click: ActivateScreen("St_Quantity Data_2", 0)
   Button "Button_5" at 163,46 size 147x30; TextOff 'Current Shift Data Minus 3'
      on Click: ActivateScreen("St_Quantity Data_3", 0)
   Button "Button_6" at 163,80 size 147x30; TextOff 'Current Shift Data Minus 4'
      on Click: ActivateScreen("St_Quantity Data_4", 0)
   Button "Button_7" at 163,113 size 147x30; TextOff 'Current Shift Data Minus 5'
      on Click: ActivateScreen("St_Quantity Data_5", 0)
   TextField "Text field_1" at 99,4 size 106x18; Text 'STATISTIC DATA'
   Button "Button_8" at 89,210 size 132x30; TextOff 'Back to Main Page'
      on Click: ActivateScreen("Main Page", 0)

